REGION Network 1
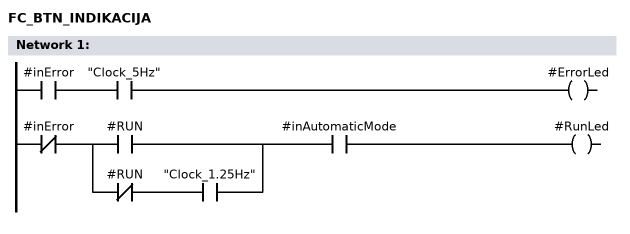
   RUNG wire#powerrail
      Contact( #inError )
      Contact( "Clock_5Hz" )
      Coil( #ErrorLed )
   END_RUNG
   RUNG wire#powerrail
      I_Contact( #inError )
      wire#w1
      Contact( #RUN )
      wire#w2
      Contact( #inAutomaticMode )
      Coil( #RunLed )
   END_RUNG
   RUNG wire#w1
      I_Contact( #RUN )
      Contact( "Clock_1.25Hz" )
   END_RUNG wire#w2
   // the same network as SCL:
   #ErrorLed := #inError AND "Clock_5Hz";
   #RunLed := NOT #inError AND (#RUN OR (NOT #RUN AND "Clock_1.25Hz")) AND #inAutomaticMode;
END_REGION
END_FUNCTION

FUNCTION "FC_SHIFT_ARRAY" : Void   // FC4, LAD
{ S7_Optimized_Access := 'TRUE' }
VERSION : 0.1
   VAR_INPUT
      InputArray : Array[0..7] of Byte;
   END_VAR
   VAR_OUTPUT
      OutputArray : Array[0..7] of Byte;
   END_VAR
   VAR_TEMP
      i : Byte;
   END_VAR
BEGIN

REGION Network 1
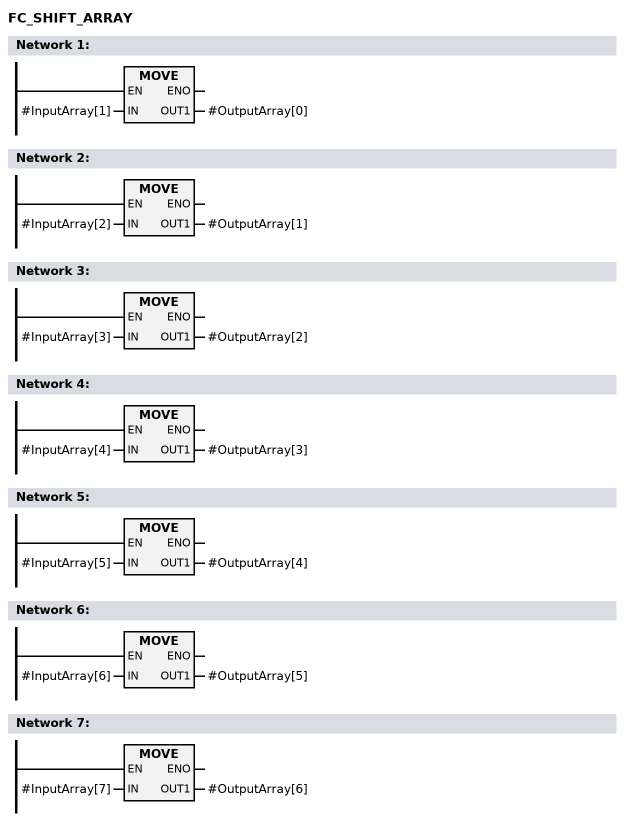
   RUNG wire#powerrail
      Move(in := #InputArray[1], out1 => #OutputArray[0])
   END_RUNG
   // the same network as SCL:
   #OutputArray[0] := #InputArray[1];
END_REGION

REGION Network 2
   RUNG wire#powerrail
      Move(in := #InputArray[2], out1 => #OutputArray[1])
   END_RUNG
   // the same network as SCL:
   #OutputArray[1] := #InputArray[2];
END_REGION

REGION Network 3
   RUNG wire#powerrail
      Move(in := #InputArray[3], out1 => #OutputArray[2])
   END_RUNG
   // the same network as SCL:
   #OutputArray[2] := #InputArray[3];
END_REGION

REGION Network 4
   RUNG wire#powerrail
      Move(in := #InputArray[4], out1 => #OutputArray[3])
   END_RUNG
   // the same network as SCL:
   #OutputArray[3] := #InputArray[4];
END_REGION

REGION Network 5
   RUNG wire#powerrail
      Move(in := #InputArray[5], out1 => #OutputArray[4])
   END_RUNG
   // the same network as SCL:
   #OutputArray[4] := #InputArray[5];
END_REGION

REGION Network 6
   RUNG wire#powerrail
      Move(in := #InputArray[6], out1 => #OutputArray[5])
   END_RUNG
   // the same network as SCL:
   #OutputArray[5] := #InputArray[6];
END_REGION

REGION Network 7
   RUNG wire#powerrail
      Move(in := #InputArray[7], out1 => #OutputArray[6])
   END_RUNG
   // the same network as SCL:
   #OutputArray[6] := #InputArray[7];
END_REGION
END_FUNCTION

ORGANIZATION_BLOCK "Main"   // OB1, LAD, ProgramCycle
TITLE = "Main Program Sweep (Cycle)"
{ S7_Optimized_Access := 'TRUE' }
VERSION : 0.1
   VAR_INPUT
      Initial_Call : Bool;   // Initial call of this OB
      Remanence : Bool;   // =True, if remanent data are available
   END_VAR
   VAR_TEMP
      stop_cikla : Bool;
      STOP_AVTO : Bool;
      temp1 : Real;
   END_VAR
   VAR_TEMP   // added for the SCL form of the ladder/FBD networks
      _w1 : Bool;
      _w2 : Bool;
      _w3 : Bool;
      _w4 : Bool;
      _w5 : Bool;
   END_VAR
BEGIN

REGION Network 1: Zagon sistema -> testiranje profinet naprav
   // testiranje io naprav
   // vklop zaslona če je OK
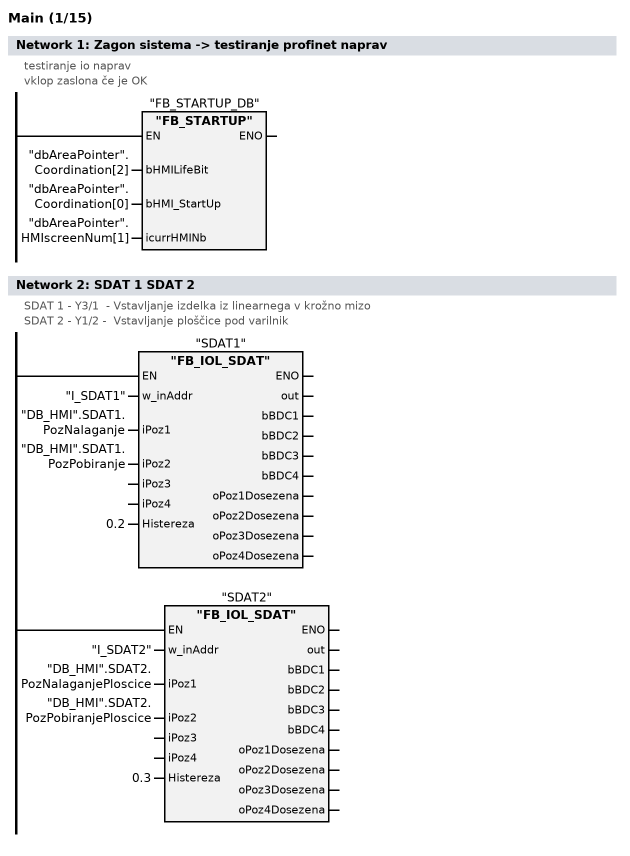
   RUNG wire#powerrail
      "FB_STARTUP_DB"(bHMILifeBit := "dbAreaPointer".Coordination[2], bHMI_StartUp := "dbAreaPointer".Coordination[0], icurrHMINb := "dbAreaPointer".HMIscreenNum[1])
   END_RUNG
   // the same network as SCL:
   "FB_STARTUP_DB"(bHMILifeBit := "dbAreaPointer".Coordination[2],   // "FB_STARTUP"
                   bHMI_StartUp := "dbAreaPointer".Coordination[0],
                   icurrHMINb := "dbAreaPointer".HMIscreenNum[1]);
END_REGION

REGION Network 2: SDAT 1 SDAT 2
   // SDAT 1 - Y3/1  - Vstavljanje izdelka iz linearnega v krožno mizo
   // SDAT 2 - Y1/2 -  Vstavljanje ploščice pod varilnik
   RUNG wire#powerrail
      "SDAT1"(w_inAddr := "I_SDAT1", iPoz1 := "DB_HMI".SDAT1.PozNalaganje, iPoz2 := "DB_HMI".SDAT1.PozPobiranje, iPoz3 :=, iPoz4 :=, Histereza := 0.2, out =>, bBDC1 =>, bBDC2 =>, bBDC3 =>, bBDC4 =>, oPoz1Dosezena =>, oPoz2Dosezena =>, oPoz3Dosezena =>, oPoz4Dosezena =>)
   END_RUNG
   RUNG wire#powerrail
      "SDAT2"(w_inAddr := "I_SDAT2", iPoz1 := "DB_HMI".SDAT2.PozNalaganjePloscice, iPoz2 := "DB_HMI".SDAT2.PozPobiranjePloscice, iPoz3 :=, iPoz4 :=, Histereza := 0.3, out =>, bBDC1 =>, bBDC2 =>, bBDC3 =>, bBDC4 =>, oPoz1Dosezena =>, oPoz2Dosezena =>, oPoz3Dosezena =>, oPoz4Dosezena =>)
   END_RUNG
   // the same network as SCL:
   "SDAT1"(w_inAddr := "I_SDAT1",   // "FB_IOL_SDAT"
           iPoz1 := "DB_HMI".SDAT1.PozNalaganje,
           iPoz2 := "DB_HMI".SDAT1.PozPobiranje,
           Histereza := 0.2);
   "SDAT2"(w_inAddr := "I_SDAT2",   // "FB_IOL_SDAT"
           iPoz1 := "DB_HMI".SDAT2.PozNalaganjePloscice,
           iPoz2 := "DB_HMI".SDAT2.PozPobiranjePloscice,
           Histereza := 0.3);
END_REGION

REGION Network 3: KEYENCE - meritve odmikov
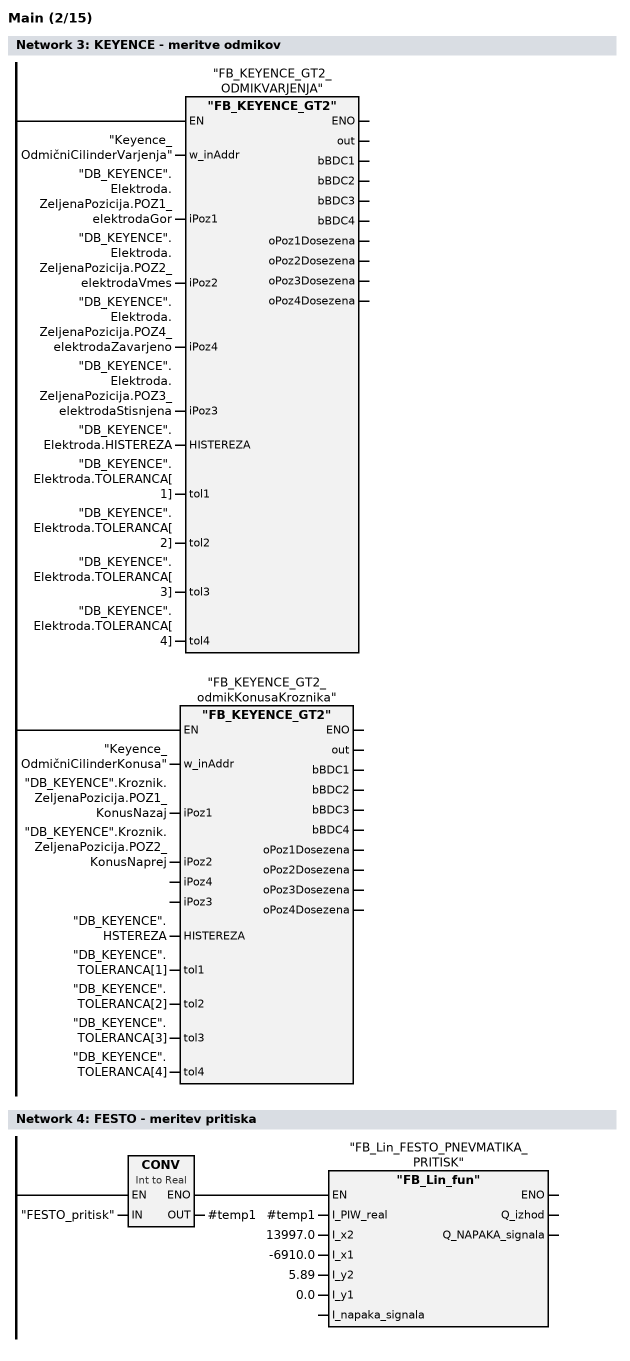
   RUNG wire#powerrail
      "FB_KEYENCE_GT2_ODMIKVARJENJA"(w_inAddr := "Keyence_OdmičniCilinderVarjenja", iPoz1 := "DB_KEYENCE".Elektroda.ZeljenaPozicija.POZ1_elektrodaGor, iPoz2 := "DB_KEYENCE".Elektroda.ZeljenaPozicija.POZ2_elektrodaVmes, iPoz4 := "DB_KEYENCE".Elektroda.ZeljenaPozicija.POZ4_elektrodaZavarjeno, iPoz3 := "DB_KEYENCE".Elektroda.ZeljenaPozicija.POZ3_elektrodaStisnjena, HISTEREZA := "DB_KEYENCE".Elektroda.HISTEREZA, tol1 := "DB_KEYENCE".Elektroda.TOLERANCA[1], tol2 := "DB_KEYENCE".Elektroda.TOLERANCA[2], tol3 := "DB_KEYENCE".Elektroda.TOLERANCA[3], tol4 := "DB_KEYENCE".Elektroda.TOLERANCA[4], out =>, bBDC1 =>, bBDC2 =>, bBDC3 =>, bBDC4 =>, oPoz1Dosezena =>, oPoz2Dosezena =>, oPoz3Dosezena =>, oPoz4Dosezena =>)
   END_RUNG
   RUNG wire#powerrail
      "FB_KEYENCE_GT2_odmikKonusaKroznika"(w_inAddr := "Keyence_OdmičniCilinderKonusa", iPoz1 := "DB_KEYENCE".Kroznik.ZeljenaPozicija.POZ1_KonusNazaj, iPoz2 := "DB_KEYENCE".Kroznik.ZeljenaPozicija.POZ2_KonusNaprej, iPoz4 :=, iPoz3 :=, HISTEREZA := "DB_KEYENCE".HSTEREZA, tol1 := "DB_KEYENCE".TOLERANCA[1], tol2 := "DB_KEYENCE".TOLERANCA[2], tol3 := "DB_KEYENCE".TOLERANCA[3], tol4 := "DB_KEYENCE".TOLERANCA[4], out =>, bBDC1 =>, bBDC2 =>, bBDC3 =>, bBDC4 =>, oPoz1Dosezena =>, oPoz2Dosezena =>, oPoz3Dosezena =>, oPoz4Dosezena =>)
   END_RUNG
   // the same network as SCL:
   "FB_KEYENCE_GT2_ODMIKVARJENJA"(w_inAddr := "Keyence_OdmičniCilinderVarjenja",   // "FB_KEYENCE_GT2"
                           iPoz1 := "DB_KEYENCE".Elektroda.ZeljenaPozicija.POZ1_elektrodaGor,
                           iPoz2 := "DB_KEYENCE".Elektroda.ZeljenaPozicija.POZ2_elektrodaVmes,
                           iPoz4 := "DB_KEYENCE".Elektroda.ZeljenaPozicija.POZ4_elektrodaZavarjeno,
                           iPoz3 := "DB_KEYENCE".Elektroda.ZeljenaPozicija.POZ3_elektrodaStisnjena,
                           HISTEREZA := "DB_KEYENCE".Elektroda.HISTEREZA,
                           tol1 := "DB_KEYENCE".Elektroda.TOLERANCA[1],
                           tol2 := "DB_KEYENCE".Elektroda.TOLERANCA[2],
                           tol3 := "DB_KEYENCE".Elektroda.TOLERANCA[3],
                           tol4 := "DB_KEYENCE".Elektroda.TOLERANCA[4]);
   "FB_KEYENCE_GT2_odmikKonusaKroznika"(w_inAddr := "Keyence_OdmičniCilinderKonusa",   // "FB_KEYENCE_GT2"
                           iPoz1 := "DB_KEYENCE".Kroznik.ZeljenaPozicija.POZ1_KonusNazaj,
                           iPoz2 := "DB_KEYENCE".Kroznik.ZeljenaPozicija.POZ2_KonusNaprej,
                           HISTEREZA := "DB_KEYENCE".HSTEREZA,
                           tol1 := "DB_KEYENCE".TOLERANCA[1],
                           tol2 := "DB_KEYENCE".TOLERANCA[2],
                           tol3 := "DB_KEYENCE".TOLERANCA[3],
                           tol4 := "DB_KEYENCE".TOLERANCA[4]);
END_REGION

REGION Network 4: FESTO - meritev pritiska
   RUNG wire#powerrail
      { S7_Templates := "[SrcType := Int, DestType := Real]" } Convert(in := "FESTO_pritisk", out => #temp1)
      "FB_Lin_FESTO_PNEVMATIKA_PRITISK"(I_PIW_real := #temp1, I_x2 := 13997.0, I_x1 := -6910.0, I_y2 := 5.89, I_y1 := 0.0, I_napaka_signala :=, Q_izhod =>, Q_NAPAKA_signala =>)
   END_RUNG
   // the same network as SCL:
   #temp1 := INT_TO_REAL("FESTO_pritisk");
   "FB_Lin_FESTO_PNEVMATIKA_PRITISK"(I_PIW_real := #temp1,   // "FB_Lin_fun"
                           I_x2 := 13997.0,
                           I_x1 := -6910.0,
                           I_y2 := 5.89,
                           I_y1 := 0.0);
END_REGION

REGION Network 5: IFM SV - Meritev pretoka & temperature
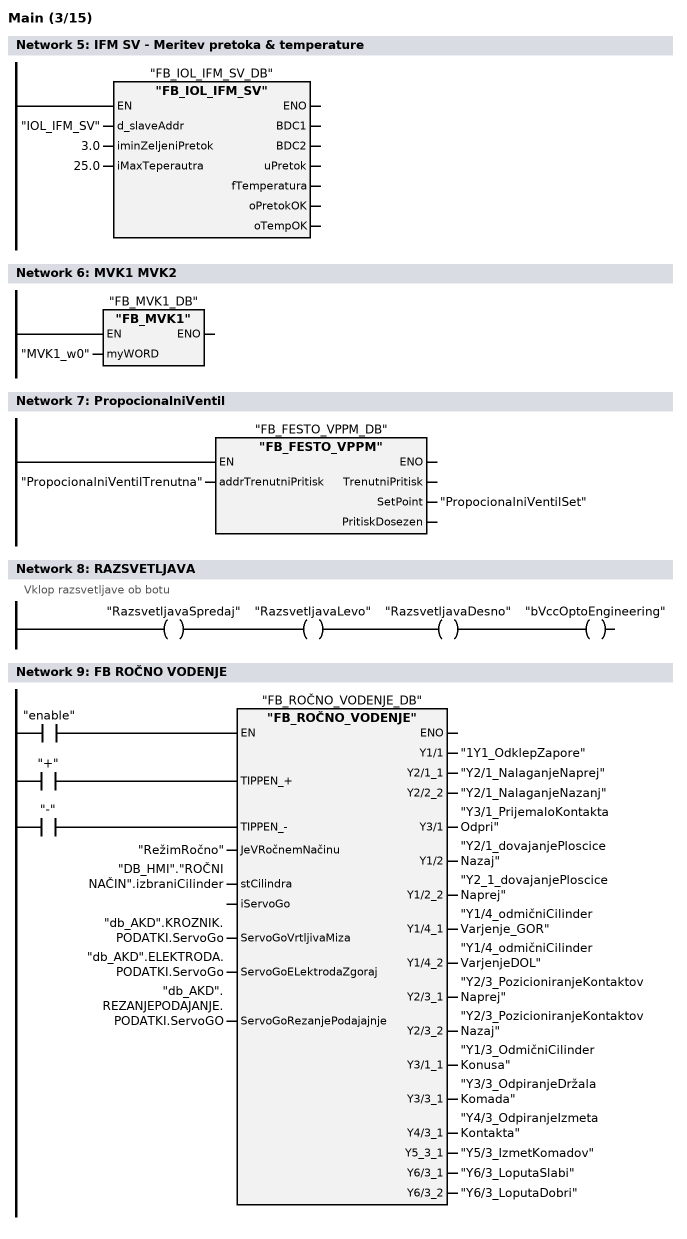
   RUNG wire#powerrail
      "FB_IOL_IFM_SV_DB"(d_slaveAddr := "IOL_IFM_SV", iminZeljeniPretok := 3.0, iMaxTeperautra := 25.0, BDC1 =>, BDC2 =>, uPretok =>, fTemperatura =>, oPretokOK =>, oTempOK =>)
   END_RUNG
   // the same network as SCL:
   "FB_IOL_IFM_SV_DB"(d_slaveAddr := "IOL_IFM_SV", iminZeljeniPretok := 3.0, iMaxTeperautra := 25.0);   // "FB_IOL_IFM_SV"
END_REGION

REGION Network 6: MVK1 MVK2
   RUNG wire#powerrail
      "FB_MVK1_DB"(myWORD := "MVK1_w0")
   END_RUNG
   // the same network as SCL:
   "FB_MVK1_DB"(myWORD := "MVK1_w0");   // "FB_MVK1"
END_REGION

REGION Network 7: PropocionalniVentil
   RUNG wire#powerrail
      "FB_FESTO_VPPM_DB"(addrTrenutniPritisk := "PropocionalniVentilTrenutna", TrenutniPritisk =>, SetPoint => "PropocionalniVentilSet", PritiskDosezen =>)
   END_RUNG
   // the same network as SCL:
   "FB_FESTO_VPPM_DB"(addrTrenutniPritisk := "PropocionalniVentilTrenutna",   // "FB_FESTO_VPPM"
                      SetPoint => "PropocionalniVentilSet");
END_REGION

REGION Network 8: RAZSVETLJAVA
   // Vklop razsvetljave ob botu
   RUNG wire#powerrail
      Coil( "RazsvetljavaSpredaj" )
      Coil( "RazsvetljavaLevo" )
      Coil( "RazsvetljavaDesno" )
      Coil( "bVccOptoEngineering" )
   END_RUNG
   // the same network as SCL:
   "RazsvetljavaSpredaj" := TRUE;
   "RazsvetljavaLevo" := TRUE;
   "RazsvetljavaDesno" := TRUE;
   "bVccOptoEngineering" := TRUE;
END_REGION

REGION Network 9: FB ROČNO VODENJE
   RUNG wire#powerrail
      Contact( "enable" )
      "FB_ROČNO_VODENJE_DB"("TIPPEN_+" := wire#w1, "TIPPEN_-" := wire#w2, JeVRočnemNačinu := "RežimRočno", stCilindra := "DB_HMI"."ROČNI NAČIN".izbraniCilinder, iServoGo :=, ServoGoVrtljivaMiza := "db_AKD".KROZNIK.PODATKI.ServoGo, ServoGoELektrodaZgoraj := "db_AKD".ELEKTRODA.PODATKI.ServoGo, ServoGoRezanjePodajajnje := "db_AKD".REZANJEPODAJANJE.PODATKI.ServoGO, "Y1/1" => "1Y1_OdklepZapore", "Y2/1_1" => "Y2/1_NalaganjeNaprej", "Y2/2_2" => "Y2/1_NalaganjeNazanj", "Y3/1" => "Y3/1_PrijemaloKontaktaOdpri", "Y1/2" => "Y2/1_dovajanjePlosciceNazaj", "Y1/2_2" => "Y2_1_dovajanjePlosciceNaprej", "Y1/4_1" => "Y1/4_odmičniCilinderVarjenje_GOR", "Y1/4_2" => "Y1/4_odmičniCilinderVarjenjeDOL", "Y2/3_1" => "Y2/3_PozicioniranjeKontaktovNaprej", "Y2/3_2" => "Y2/3_PozicioniranjeKontaktovNazaj", "Y3/1_1" => "Y1/3_OdmičniCilinderKonusa", "Y3/3_1" => "Y3/3_OdpiranjeDržalaKomada", "Y4/3_1" => "Y4/3_OdpiranjeIzmetaKontakta", Y5_3_1 => "Y5/3_IzmetKomadov", "Y6/3_1" => "Y6/3_LoputaSlabi", "Y6/3_2" => "Y6/3_LoputaDobri")
   END_RUNG
   RUNG wire#powerrail
      Contact( "+" )
   END_RUNG wire#w1
   RUNG wire#powerrail
      Contact( "-" )
   END_RUNG wire#w2
   // the same network as SCL:
   IF "enable" THEN
       "FB_ROČNO_VODENJE_DB"("TIPPEN_+" := "+",   // "FB_ROČNO_VODENJE"
                             "TIPPEN_-" := "-",
                             JeVRočnemNačinu := "RežimRočno",
                             stCilindra := "DB_HMI"."ROČNI NAČIN".izbraniCilinder,
                             ServoGoVrtljivaMiza := "db_AKD".KROZNIK.PODATKI.ServoGo,
                             ServoGoELektrodaZgoraj := "db_AKD".ELEKTRODA.PODATKI.ServoGo,
                             ServoGoRezanjePodajajnje := "db_AKD".REZANJEPODAJANJE.PODATKI.ServoGO,
                             "Y1/1" => "1Y1_OdklepZapore",
                             "Y2/1_1" => "Y2/1_NalaganjeNaprej",
                             "Y2/2_2" => "Y2/1_NalaganjeNazanj",
                             "Y3/1" => "Y3/1_PrijemaloKontaktaOdpri",
                             "Y1/2" => "Y2/1_dovajanjePlosciceNazaj",
                             "Y1/2_2" => "Y2_1_dovajanjePlosciceNaprej",
                             "Y1/4_1" => "Y1/4_odmičniCilinderVarjenje_GOR",
                             "Y1/4_2" => "Y1/4_odmičniCilinderVarjenjeDOL",
                             "Y2/3_1" => "Y2/3_PozicioniranjeKontaktovNaprej",
                             "Y2/3_2" => "Y2/3_PozicioniranjeKontaktovNazaj",
                             "Y3/1_1" => "Y1/3_OdmičniCilinderKonusa",
                             "Y3/3_1" => "Y3/3_OdpiranjeDržalaKomada",
                             "Y4/3_1" => "Y4/3_OdpiranjeIzmetaKontakta",
                             Y5_3_1 => "Y5/3_IzmetKomadov",
                             "Y6/3_1" => "Y6/3_LoputaSlabi",
                             "Y6/3_2" => "Y6/3_LoputaDobri");
   END_IF;
END_REGION

REGION Network 10: GL program - SEQ
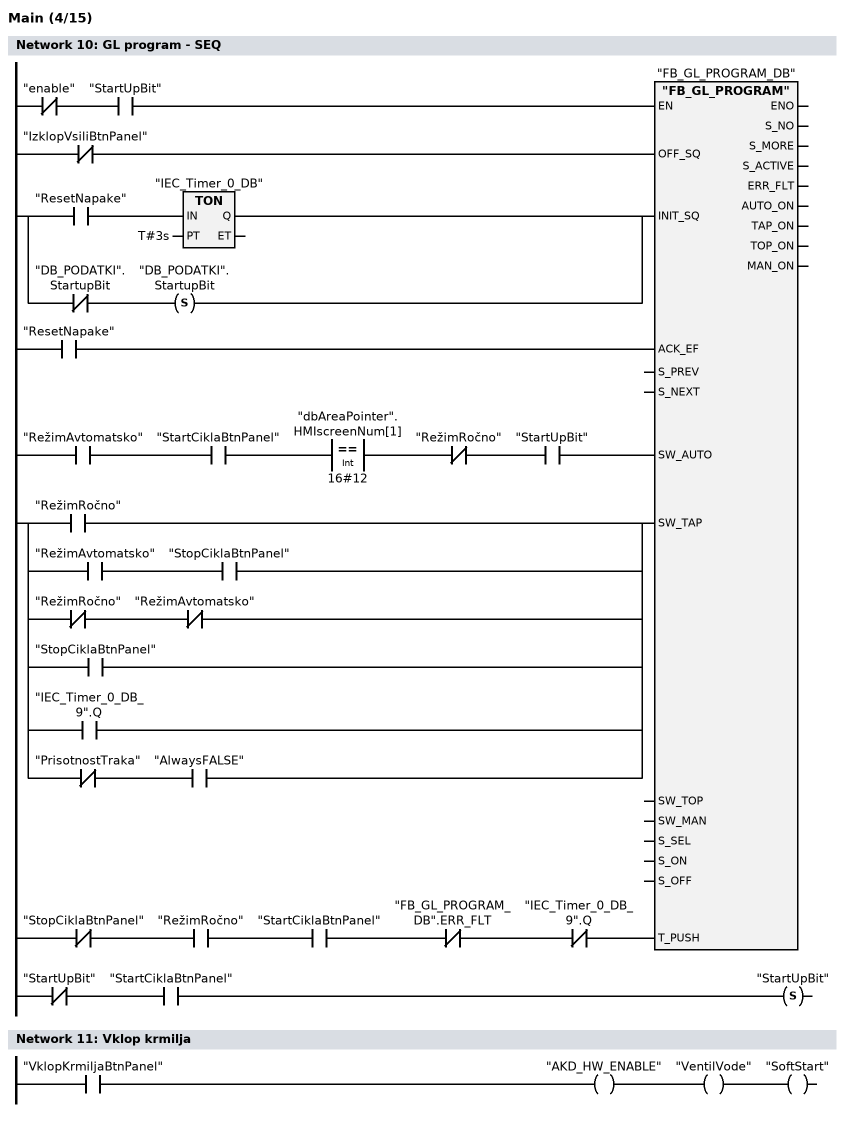
   "IEC_Timer_0_DB".TON(IN := "ResetNapake", PT := T#3s);
   #_w1 := NOT "DB_PODATKI".StartupBit;
   IF #_w1 THEN "DB_PODATKI".StartupBit := TRUE; END_IF;
   IF NOT "enable" AND "StartUpBit" THEN
       "FB_GL_PROGRAM_DB"(OFF_SQ := NOT "IzklopVsiliBtnPanel",   // "FB_GL_PROGRAM"
                          INIT_SQ := "IEC_Timer_0_DB".Q OR #_w1,
                          ACK_EF := "ResetNapake",
                          SW_AUTO := "RežimAvtomatsko" AND "StartCiklaBtnPanel" AND ("dbAreaPointer".HMIscreenNum[1] = 16#12) AND NOT "RežimRočno" AND "StartUpBit",
                          SW_TAP := "RežimRočno" OR ("RežimAvtomatsko" AND "StopCiklaBtnPanel") OR (NOT "RežimRočno" AND NOT "RežimAvtomatsko") OR "StopCiklaBtnPanel" OR "IEC_Timer_0_DB_9".Q OR (NOT "PrisotnostTraka" AND "AlwaysFALSE"),
                          T_PUSH := NOT "StopCiklaBtnPanel" AND "RežimRočno" AND "StartCiklaBtnPanel" AND NOT "FB_GL_PROGRAM_DB".ERR_FLT AND NOT "IEC_Timer_0_DB_9".Q);
   END_IF;
   IF NOT "StartUpBit" AND "StartCiklaBtnPanel" THEN "StartUpBit" := TRUE; END_IF;
END_REGION

REGION Network 11: Vklop krmilja
   RUNG wire#powerrail
      Contact( "VklopKrmiljaBtnPanel" )
      Coil( "AKD_HW_ENABLE" )
      Coil( "VentilVode" )
      Coil( "SoftStart" )
   END_RUNG
   // the same network as SCL:
   "AKD_HW_ENABLE" := "VklopKrmiljaBtnPanel";
   "VentilVode" := "VklopKrmiljaBtnPanel";
   "SoftStart" := "VklopKrmiljaBtnPanel";
END_REGION

REGION Network 12: PREKLOP HMI - ROČNO <> AVTO
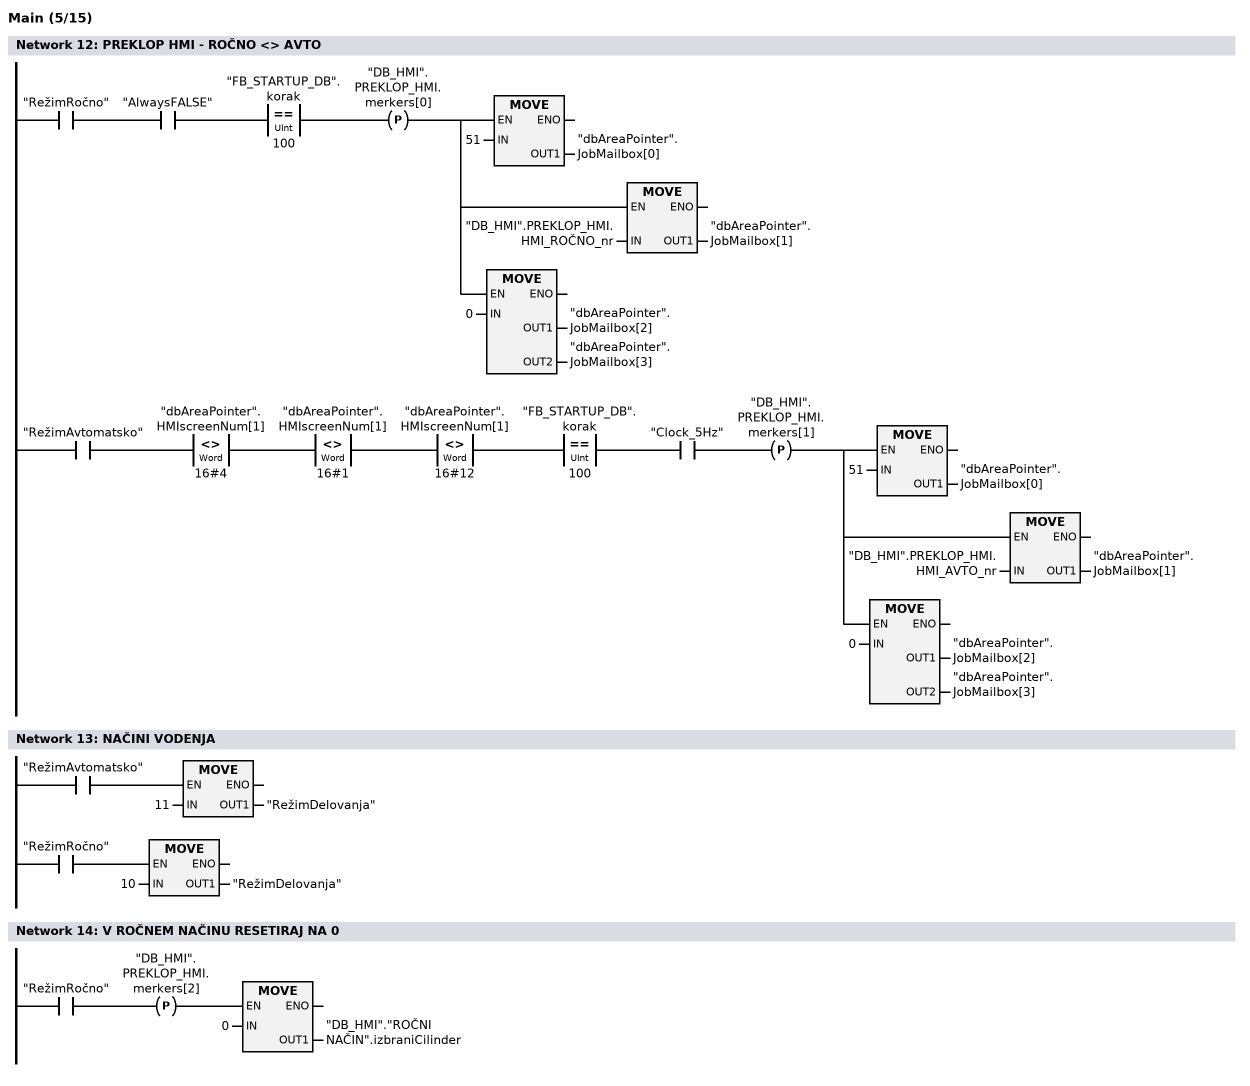
   RUNG wire#powerrail
      Contact( "RežimRočno" )
      Contact( "AlwaysFALSE" )
      { S7_Templates := "SrcType := UInt" } EQ_Contact(in1 := "FB_STARTUP_DB".korak, in2 := 100)
      P_Trig( "DB_HMI".PREKLOP_HMI.merkers[0] )
      wire#w1
      Move(in := 51, out1 => "dbAreaPointer".JobMailbox[0])
   END_RUNG
   RUNG wire#w1
      Move(in := "DB_HMI".PREKLOP_HMI.HMI_ROČNO_nr, out1 => "dbAreaPointer".JobMailbox[1])
   END_RUNG
   RUNG wire#w1
      Move(in := 0, out1 => "dbAreaPointer".JobMailbox[2], out2 => "dbAreaPointer".JobMailbox[3])
   END_RUNG
   RUNG wire#powerrail
      Contact( "RežimAvtomatsko" )
      { S7_Templates := "SrcType := Word" } NE_Contact(in1 := "dbAreaPointer".HMIscreenNum[1], in2 := 16#4)
      { S7_Templates := "SrcType := Word" } NE_Contact(in1 := "dbAreaPointer".HMIscreenNum[1], in2 := 16#1)
      { S7_Templates := "SrcType := Word" } NE_Contact(in1 := "dbAreaPointer".HMIscreenNum[1], in2 := 16#12)
      { S7_Templates := "SrcType := UInt" } EQ_Contact(in1 := "FB_STARTUP_DB".korak, in2 := 100)
      Contact( "Clock_5Hz" )
      P_Trig( "DB_HMI".PREKLOP_HMI.merkers[1] )
      wire#w2
      Move(in := 51, out1 => "dbAreaPointer".JobMailbox[0])
   END_RUNG
   RUNG wire#w2
      Move(in := "DB_HMI".PREKLOP_HMI.HMI_AVTO_nr, out1 => "dbAreaPointer".JobMailbox[1])
   END_RUNG
   RUNG wire#w2
      Move(in := 0, out1 => "dbAreaPointer".JobMailbox[2], out2 => "dbAreaPointer".JobMailbox[3])
   END_RUNG
   // the same network as SCL:
   #_w1 := "RežimRočno" AND "AlwaysFALSE" AND ("FB_STARTUP_DB".korak = 100);
   #_w2 := #_w1 AND NOT "DB_HMI".PREKLOP_HMI.merkers[0];   // rising edge
   "DB_HMI".PREKLOP_HMI.merkers[0] := #_w1;
   IF #_w2 THEN
       "dbAreaPointer".JobMailbox[0] := 51;
       "dbAreaPointer".JobMailbox[1] := "DB_HMI".PREKLOP_HMI.HMI_ROČNO_nr;
       "dbAreaPointer".JobMailbox[2] := 0;
       "dbAreaPointer".JobMailbox[3] := 0;
   END_IF;
   #_w3 := "RežimAvtomatsko" AND ("dbAreaPointer".HMIscreenNum[1] <> 16#4) AND ("dbAreaPointer".HMIscreenNum[1] <> 16#1) AND ("dbAreaPointer".HMIscreenNum[1] <> 16#12) AND ("FB_STARTUP_DB".korak = 100) AND "Clock_5Hz";
   #_w4 := #_w3 AND NOT "DB_HMI".PREKLOP_HMI.merkers[1];   // rising edge
   "DB_HMI".PREKLOP_HMI.merkers[1] := #_w3;
   IF #_w4 THEN
       "dbAreaPointer".JobMailbox[0] := 51;
       "dbAreaPointer".JobMailbox[1] := "DB_HMI".PREKLOP_HMI.HMI_AVTO_nr;
       "dbAreaPointer".JobMailbox[2] := 0;
       "dbAreaPointer".JobMailbox[3] := 0;
   END_IF;
END_REGION

REGION Network 13: NAČINI VODENJA
   RUNG wire#powerrail
      Contact( "RežimAvtomatsko" )
      Move(in := 11, out1 => "RežimDelovanja")
   END_RUNG
   RUNG wire#powerrail
      Contact( "RežimRočno" )
      Move(in := 10, out1 => "RežimDelovanja")
   END_RUNG
   // the same network as SCL:
   IF "RežimAvtomatsko" THEN "RežimDelovanja" := 11; END_IF;
   IF "RežimRočno" THEN "RežimDelovanja" := 10; END_IF;
END_REGION

REGION Network 14: V ROČNEM NAČINU RESETIRAJ NA 0
   RUNG wire#powerrail
      Contact( "RežimRočno" )
      P_Trig( "DB_HMI".PREKLOP_HMI.merkers[2] )
      Move(in := 0, out1 => "DB_HMI"."ROČNI NAČIN".izbraniCilinder)
   END_RUNG
   // the same network as SCL:
   #_w1 := "RežimRočno" AND NOT "DB_HMI".PREKLOP_HMI.merkers[2];   // rising edge
   "DB_HMI".PREKLOP_HMI.merkers[2] := "RežimRočno";
   IF #_w1 THEN "DB_HMI"."ROČNI NAČIN".izbraniCilinder := 0; END_IF;
END_REGION

REGION Network 15: UDP komunikacija - Izklop PCja - TUSEND
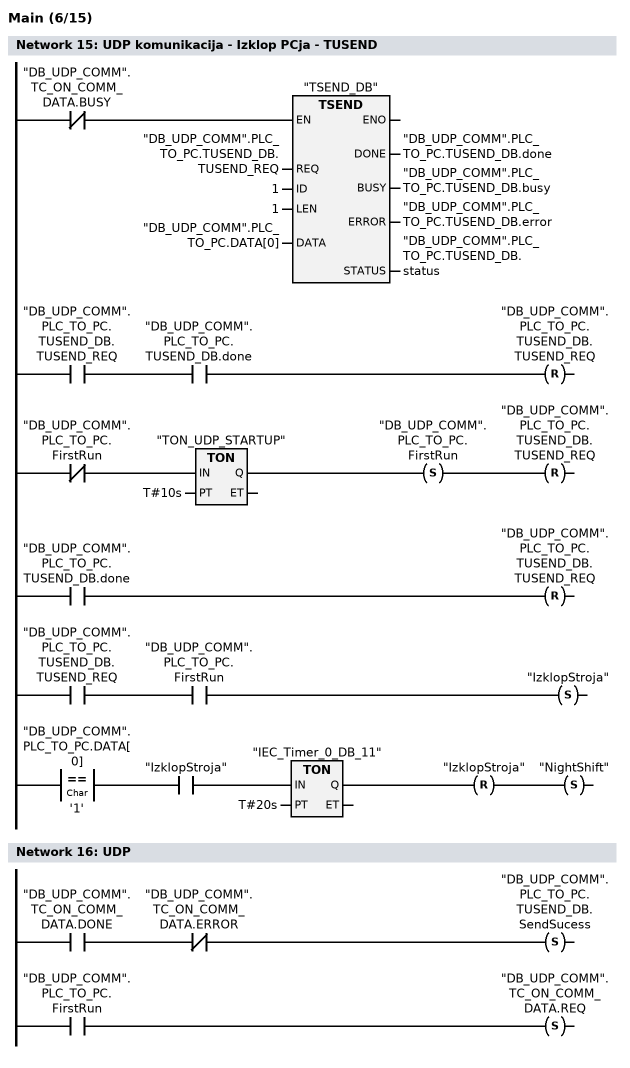
   IF NOT "DB_UDP_COMM".TC_ON_COMM_DATA.BUSY THEN
       "TSEND_DB"(REQ := "DB_UDP_COMM".PLC_TO_PC.TUSEND_DB.TUSEND_REQ,   // TSEND
                  ID := 1,
                  LEN := 1,
                  DATA := "DB_UDP_COMM".PLC_TO_PC.DATA[0],
                  DONE => "DB_UDP_COMM".PLC_TO_PC.TUSEND_DB.done,
                  BUSY => "DB_UDP_COMM".PLC_TO_PC.TUSEND_DB.busy,
                  ERROR => "DB_UDP_COMM".PLC_TO_PC.TUSEND_DB.error,
                  STATUS => "DB_UDP_COMM".PLC_TO_PC.TUSEND_DB.status);
   END_IF;
   IF "DB_UDP_COMM".PLC_TO_PC.TUSEND_DB.TUSEND_REQ AND "DB_UDP_COMM".PLC_TO_PC.TUSEND_DB.done THEN
       "DB_UDP_COMM".PLC_TO_PC.TUSEND_DB.TUSEND_REQ := FALSE;
   END_IF;
   "TON_UDP_STARTUP".TON(IN := NOT "DB_UDP_COMM".PLC_TO_PC.FirstRun, PT := T#10s);
   IF "TON_UDP_STARTUP".Q THEN
       "DB_UDP_COMM".PLC_TO_PC.FirstRun := TRUE;
       "DB_UDP_COMM".PLC_TO_PC.TUSEND_DB.TUSEND_REQ := FALSE;
   END_IF;
   IF "DB_UDP_COMM".PLC_TO_PC.TUSEND_DB.done THEN
       "DB_UDP_COMM".PLC_TO_PC.TUSEND_DB.TUSEND_REQ := FALSE;
   END_IF;
   IF "DB_UDP_COMM".PLC_TO_PC.TUSEND_DB.TUSEND_REQ AND "DB_UDP_COMM".PLC_TO_PC.FirstRun THEN
       "IzklopStroja" := TRUE;
   END_IF;
   "IEC_Timer_0_DB_11".TON(IN := ("DB_UDP_COMM".PLC_TO_PC.DATA[0] = '1') AND "IzklopStroja", PT := T#20s);
   IF "IEC_Timer_0_DB_11".Q THEN
       "IzklopStroja" := FALSE;
       "NightShift" := TRUE;
   END_IF;
END_REGION

REGION Network 16: UDP
   RUNG wire#powerrail
      Contact( "DB_UDP_COMM".TC_ON_COMM_DATA.DONE )
      I_Contact( "DB_UDP_COMM".TC_ON_COMM_DATA.ERROR )
      S_Coil( "DB_UDP_COMM".PLC_TO_PC.TUSEND_DB.SendSucess )
   END_RUNG
   RUNG wire#powerrail
      Contact( "DB_UDP_COMM".PLC_TO_PC.FirstRun )
      S_Coil( "DB_UDP_COMM".TC_ON_COMM_DATA.REQ )
   END_RUNG
   // the same network as SCL:
   IF "DB_UDP_COMM".TC_ON_COMM_DATA.DONE AND NOT "DB_UDP_COMM".TC_ON_COMM_DATA.ERROR THEN
       "DB_UDP_COMM".PLC_TO_PC.TUSEND_DB.SendSucess := TRUE;
   END_IF;
   IF "DB_UDP_COMM".PLC_TO_PC.FirstRun THEN "DB_UDP_COMM".TC_ON_COMM_DATA.REQ := TRUE; END_IF;
END_REGION

REGION Network 17: UDP TCON